   "DB_MouldEditor_HMI_uData_arShotSet{0}_Pressure{4}" : Real = PLC DB_MouldEditor_HMI.uData.arShotSet[0].Pressure[4] AT %DB10.DBD126, 1 s
   "DB_MouldEditor_HMI_uData_arShotSet{0}_Pressure{5}" : Real = PLC DB_MouldEditor_HMI.uData.arShotSet[0].Pressure[5] AT %DB10.DBD130, 1 s
   "DB_MouldEditor_HMI_uData_arShotSet{0}_Pressure{6}" : Real = PLC DB_MouldEditor_HMI.uData.arShotSet[0].Pressure[6] AT %DB10.DBD134, 1 s
   "DB_MouldEditor_HMI_uData_arShotSet{0}_Flow{1}" : Real = PLC DB_MouldEditor_HMI.uData.arShotSet[0].Flow[1] AT %DB10.DBD138, 1 s
   "DB_MouldEditor_HMI_uData_arShotSet{0}_Flow{2}" : Real = PLC DB_MouldEditor_HMI.uData.arShotSet[0].Flow[2] AT %DB10.DBD142, 1 s
   "DB_MouldEditor_HMI_uData_arShotSet{0}_Flow{3}" : Real = PLC DB_MouldEditor_HMI.uData.arShotSet[0].Flow[3] AT %DB10.DBD146, 1 s
   "DB_MouldEditor_HMI_uData_arShotSet{0}_Flow{4}" : Real = PLC DB_MouldEditor_HMI.uData.arShotSet[0].Flow[4] AT %DB10.DBD150, 1 s
   "DB_MouldEditor_HMI_uData_arShotSet{0}_Flow{5}" : Real = PLC DB_MouldEditor_HMI.uData.arShotSet[0].Flow[5] AT %DB10.DBD154, 1 s
   "DB_MouldEditor_HMI_uData_arShotSet{0}_Flow{6}" : Real = PLC DB_MouldEditor_HMI.uData.arShotSet[0].Flow[6] AT %DB10.DBD158, 1 s
   "DB_MouldEditor_HMI_uData_arShotSet{1}_Pressure{1}" : Real = PLC DB_MouldEditor_HMI.uData.arShotSet[1].Pressure[1] AT %DB10.DBD186, 1 s
   "DB_MouldEditor_HMI_uData_arShotSet{1}_Pressure{2}" : Real = PLC DB_MouldEditor_HMI.uData.arShotSet[1].Pressure[2] AT %DB10.DBD190, 1 s
   "DB_MouldEditor_HMI_uData_arShotSet{1}_Pressure{3}" : Real = PLC DB_MouldEditor_HMI.uData.arShotSet[1].Pressure[3] AT %DB10.DBD194, 1 s
   "DB_MouldEditor_HMI_uData_arShotSet{1}_Pressure{4}" : Real = PLC DB_MouldEditor_HMI.uData.arShotSet[1].Pressure[4] AT %DB10.DBD198, 1 s
   "DB_MouldEditor_HMI_uData_arShotSet{1}_Pressure{5}" : Real = PLC DB_MouldEditor_HMI.uData.arShotSet[1].Pressure[5] AT %DB10.DBD202, 1 s
   "DB_MouldEditor_HMI_uData_arShotSet{1}_Pressure{6}" : Real = PLC DB918_ShotResultlast10.FilteredShot[2].Mixingratio[1] AT %DB10.DBD206, 1 s
   "DB_MouldEditor_HMI_uData_arShotSet{1}_Flow{1}" : Real = PLC DB_MouldEditor_HMI.uData.arShotSet[1].Flow[1] AT %DB10.DBD210, 1 s
   "DB_MouldEditor_HMI_uData_arShotSet{1}_Flow{2}" : Real = PLC DB_MouldEditor_HMI.uData.arShotSet[1].Flow[2] AT %DB10.DBD214, 1 s
   "DB_MouldEditor_HMI_uData_arShotSet{1}_Flow{3}" : Real = PLC DB_MouldEditor_HMI.uData.arShotSet[1].Flow[3] AT %DB10.DBD218, 1 s
   "DB_MouldEditor_HMI_uData_arShotSet{1}_Flow{4}" : Real = PLC DB_MouldEditor_HMI.uData.arShotSet[1].Flow[4] AT %DB10.DBD222, 1 s
   "DB_MouldEditor_HMI_uData_arShotSet{1}_Flow{5}" : Real = PLC DB_MouldEditor_HMI.uData.arShotSet[1].Flow[5] AT %DB10.DBD226, 1 s
   "DB_MouldEditor_HMI_uData_arShotSet{1}_Flow{6}" : Real = PLC DB_MouldEditor_HMI.uData.arShotSet[1].Flow[6] AT %DB10.DBD230, 1 s
   "DB_MouldEditor_HMI_uData_arShotSet{2}_Pressure{1}" : Real = PLC DB_MouldEditor_HMI.uData.arShotSet[2].Pressure[1] AT %DB10.DBD258, 1 s
   "DB_MouldEditor_HMI_uData_arShotSet{2}_Pressure{2}" : Real = PLC DB_MouldEditor_HMI.uData.arShotSet[2].Pressure[2] AT %DB10.DBD262, 1 s
   "DB_MouldEditor_HMI_uData_arShotSet{2}_Pressure{3}" : Real = PLC DB_MouldEditor_HMI.uData.arShotSet[2].Pressure[3] AT %DB10.DBD266, 1 s
   "DB_MouldEditor_HMI_uData_arShotSet{2}_Pressure{4}" : Real = PLC DB_MouldEditor_HMI.uData.arShotSet[2].Pressure[4] AT %DB10.DBD270, 1 s
   "DB_MouldEditor_HMI_uData_arShotSet{2}_Pressure{5}" : Real = PLC DB_MouldEditor_HMI.uData.arShotSet[2].Pressure[5] AT %DB10.DBD274, 1 s
   "DB_MouldEditor_HMI_uData_arShotSet{2}_Pressure{6}" : Real = PLC DB_MouldEditor_HMI.uData.arShotSet[2].Pressure[6] AT %DB10.DBD278, 1 s
   "DB_MouldEditor_HMI_uData_arShotSet{2}_Flow{1}" : Real = PLC DB_MouldEditor_HMI.uData.arShotSet[2].Flow[1] AT %DB10.DBD282, 1 s
   "DB_MouldEditor_HMI_uData_arShotSet{2}_Flow{2}" : Real = PLC DB_MouldEditor_HMI.uData.arShotSet[2].Flow[2] AT %DB10.DBD286, 1 s
   "DB_MouldEditor_HMI_uData_arShotSet{2}_Flow{3}" : Real = PLC DB_MouldEditor_HMI.uData.arShotSet[2].Flow[3] AT %DB10.DBD290, 1 s
   "DB_MouldEditor_HMI_uData_arShotSet{2}_Flow{4}" : Real = PLC DB_MouldEditor_HMI.uData.arShotSet[2].Flow[4] AT %DB10.DBD294, 1 s
   "DB_MouldEditor_HMI_uData_arShotSet{2}_Flow{5}" : Real = PLC DB_MouldEditor_HMI.uData.arShotSet[2].Flow[5] AT %DB10.DBD298, 1 s
   "DB_MouldEditor_HMI_uData_arShotSet{2}_Flow{6}" : Real = PLC DB_MouldEditor_HMI.uData.arShotSet[2].Flow[6] AT %DB10.DBD302, 1 s
   "DB_MouldEditor_HMI_uData_arShotSet{3}_Pressure{1}" : Real = PLC DB_MouldEditor_HMI.uData.arShotSet[3].Pressure[1] AT %DB10.DBD330, 1 s
   "DB_MouldEditor_HMI_uData_arShotSet{3}_Pressure{2}" : Real = PLC DB_MouldEditor_HMI.uData.arShotSet[3].Pressure[2] AT %DB10.DBD334, 1 s
   "DB_MouldEditor_HMI_uData_arShotSet{3}_Pressure{3}" : Real = PLC DB_MouldEditor_HMI.uData.arShotSet[3].Pressure[3] AT %DB10.DBD338, 1 s
   "DB_MouldEditor_HMI_uData_arShotSet{3}_Pressure{4}" : Real = PLC DB_MouldEditor_HMI.uData.arShotSet[3].Pressure[4] AT %DB10.DBD342, 1 s
   "DB_MouldEditor_HMI_uData_arShotSet{3}_Pressure{5}" : Real = PLC DB_MouldEditor_HMI.uData.arShotSet[3].Pressure[5] AT %DB10.DBD346, 1 s
   "DB_MouldEditor_HMI_uData_arShotSet{3}_Pressure{6}" : Real = PLC DB_MouldEditor_HMI.uData.arShotSet[3].Pressure[6] AT %DB10.DBD350, 1 s
   "DB_MouldEditor_HMI_uData_arShotSet{3}_Flow{1}" : Real = PLC DB_MouldEditor_HMI.uData.arShotSet[3].Flow[1] AT %DB10.DBD354, 1 s
   "DB_MouldEditor_HMI_uData_arShotSet{3}_Flow{2}" : Real = PLC DB_MouldEditor_HMI.uData.arShotSet[3].Flow[2] AT %DB10.DBD358, 1 s
   "DB_MouldEditor_HMI_uData_arShotSet{3}_Flow{3}" : Real = PLC DB_MouldEditor_HMI.uData.arShotSet[3].Flow[3] AT %DB10.DBD362, 1 s
   "DB_MouldEditor_HMI_uData_arShotSet{3}_Flow{4}" : Real = PLC DB_MouldEditor_HMI.uData.arShotSet[3].Flow[4] AT %DB10.DBD366, 1 s
   "DB_MouldEditor_HMI_uData_arShotSet{3}_Flow{5}" : Real = PLC DB_MouldEditor_HMI.uData.arShotSet[3].Flow[5] AT %DB10.DBD370, 1 s
   "DB_MouldEditor_HMI_uData_arShotSet{3}_Flow{6}" : Real = PLC DB_MouldEditor_HMI.uData.arShotSet[3].Flow[6] AT %DB10.DBD374, 1 s
   "DB_MouldEditor_HMI_uData_arShotSet{4}_Pressure{1}" : Real = PLC DB_MouldEditor_HMI.uData.arShotSet[4].Pressure[1] AT %DB10.DBD402, 1 s
   "DB_MouldEditor_HMI_uData_arShotSet{4}_Pressure{2}" : Real = PLC DB_MouldEditor_HMI.uData.arShotSet[4].Pressure[2] AT %DB10.DBD406, 1 s
   "DB_MouldEditor_HMI_uData_arShotSet{4}_Pressure{3}" : Real = PLC DB_MouldEditor_HMI.uData.arShotSet[4].Pressure[3] AT %DB10.DBD410, 1 s
   "DB_MouldEditor_HMI_uData_arShotSet{4}_Pressure{4}" : Real = PLC DB_MouldEditor_HMI.uData.arShotSet[4].Pressure[4] AT %DB10.DBD414, 1 s
   "DB_MouldEditor_HMI_uData_arShotSet{4}_Pressure{5}" : Real = PLC DB_MouldEditor_HMI.uData.arShotSet[4].Pressure[5] AT %DB10.DBD418, 1 s
   "DB_MouldEditor_HMI_uData_arShotSet{4}_Pressure{6}" : Real = PLC DB_MouldEditor_HMI.uData.arShotSet[4].Pressure[6] AT %DB10.DBD422, 1 s
   "DB_MouldEditor_HMI_uData_arShotSet{4}_Flow{1}" : Real = PLC DB_MouldEditor_HMI.uData.arShotSet[4].Flow[1] AT %DB10.DBD426, 1 s
   "DB_MouldEditor_HMI_uData_arShotSet{4}_Flow{2}" : Real = PLC DB_MouldEditor_HMI.uData.arShotSet[4].Flow[2] AT %DB10.DBD430, 1 s
   "DB_MouldEditor_HMI_uData_arShotSet{4}_Flow{3}" : Real = PLC DB_MouldEditor_HMI.uData.arShotSet[4].Flow[3] AT %DB10.DBD434, 1 s
   "DB_MouldEditor_HMI_uData_arShotSet{4}_Flow{4}" : Real = PLC DB_MouldEditor_HMI.uData.arShotSet[4].Flow[4] AT %DB10.DBD438, 1 s
   "DB_MouldEditor_HMI_uData_arShotSet{4}_Flow{5}" : Real = PLC DB_MouldEditor_HMI.uData.arShotSet[4].Flow[5] AT %DB10.DBD442, 1 s
   "DB_MouldEditor_HMI_uData_arShotSet{4}_Flow{6}" : Real = PLC DB_MouldEditor_HMI.uData.arShotSet[4].Flow[6] AT %DB10.DBD446, 1 s
   "DB_MouldEditor_HMI_uData_arShotSet{5}_Pressure{1}" : Real = PLC DB_MouldEditor_HMI.uData.arShotSet[5].Pressure[1] AT %DB10.DBD474, 1 s
   "DB_MouldEditor_HMI_uData_arShotSet{5}_Pressure{2}" : Real = PLC DB_MouldEditor_HMI.uData.arShotSet[5].Pressure[2] AT %DB10.DBD478, 1 s
   "DB_MouldEditor_HMI_uData_arShotSet{5}_Pressure{3}" : Real = PLC DB_MouldEditor_HMI.uData.arShotSet[5].Pressure[3] AT %DB10.DBD482, 1 s
   "DB_MouldEditor_HMI_uData_arShotSet{5}_Pressure{4}" : Real = PLC DB_MouldEditor_HMI.uData.arShotSet[5].Pressure[4] AT %DB10.DBD486, 1 s
   "DB_MouldEditor_HMI_uData_arShotSet{5}_Pressure{5}" : Real = PLC DB_MouldEditor_HMI.uData.arShotSet[5].Pressure[5] AT %DB10.DBD490, 1 s
   "DB_MouldEditor_HMI_uData_arShotSet{5}_Pressure{6}" : Real = PLC DB_MouldEditor_HMI.uData.arShotSet[5].Pressure[6] AT %DB10.DBD494, 1 s
   "DB_MouldEditor_HMI_uData_arShotSet{5}_Flow{1}" : Real = PLC DB_MouldEditor_HMI.uData.arShotSet[5].Flow[1] AT %DB10.DBD498, 1 s
   "DB_MouldEditor_HMI_uData_arShotSet{5}_Flow{2}" : Real = PLC DB_MouldEditor_HMI.uData.arShotSet[5].Flow[2] AT %DB10.DBD502, 1 s
   "DB_MouldEditor_HMI_uData_arShotSet{5}_Flow{3}" : Real = PLC DB_MouldEditor_HMI.uData.arShotSet[5].Flow[3] AT %DB10.DBD506, 1 s
   "DB_MouldEditor_HMI_uData_arShotSet{5}_Flow{4}" : Real = PLC DB_MouldEditor_HMI.uData.arShotSet[5].Flow[4] AT %DB10.DBD510, 1 s
   "DB_MouldEditor_HMI_uData_arShotSet{5}_Flow{5}" : Real = PLC DB_MouldEditor_HMI.uData.arShotSet[5].Flow[5] AT %DB10.DBD514, 1 s
   "DB_MouldEditor_HMI_uData_arShotSet{5}_Flow{6}" : Real = PLC DB_MouldEditor_HMI.uData.arShotSet[5].Flow[6] AT %DB10.DBD518, 1 s
   "DB_MouldEditor_HMI_uData_arShotSet{6}_Pressure{1}" : Real = PLC DB_MouldEditor_HMI.uData.arShotSet[6].Pressure[1] AT %DB10.DBD546, 1 s
   "DB_MouldEditor_HMI_uData_arShotSet{6}_Pressure{2}" : Real = PLC DB_MouldEditor_HMI.uData.arShotSet[6].Pressure[2] AT %DB10.DBD550, 1 s
   "DB_MouldEditor_HMI_uData_arShotSet{6}_Pressure{3}" : Real = PLC DB_MouldEditor_HMI.uData.arShotSet[6].Pressure[3] AT %DB10.DBD554, 1 s
   "DB_MouldEditor_HMI_uData_arShotSet{6}_Pressure{4}" : Real = PLC DB_MouldEditor_HMI.uData.arShotSet[6].Pressure[4] AT %DB10.DBD558, 1 s
   "DB_MouldEditor_HMI_uData_arShotSet{6}_Pressure{5}" : Real = PLC DB_MouldEditor_HMI.uData.arShotSet[6].Pressure[5] AT %DB10.DBD562, 1 s
   "DB_MouldEditor_HMI_uData_arShotSet{6}_Pressure{6}" : Real = PLC DB_MouldEditor_HMI.uData.arShotSet[6].Pressure[6] AT %DB10.DBD566, 1 s
   "DB_MouldEditor_HMI_uData_arShotSet{6}_Flow{1}" : Real = PLC DB_MouldEditor_HMI.uData.arShotSet[6].Flow[1] AT %DB10.DBD570, 1 s
   "DB_MouldEditor_HMI_uData_arShotSet{6}_Flow{2}" : Real = PLC DB_MouldEditor_HMI.uData.arShotSet[6].Flow[2] AT %DB10.DBD574, 1 s
   "DB_MouldEditor_HMI_uData_arShotSet{6}_Flow{3}" : Real = PLC DB_MouldEditor_HMI.uData.arShotSet[6].Flow[3] AT %DB10.DBD578, 1 s
   "DB_MouldEditor_HMI_uData_arShotSet{6}_Flow{4}" : Real = PLC DB_MouldEditor_HMI.uData.arShotSet[6].Flow[4] AT %DB10.DBD582, 1 s
   "DB_MouldEditor_HMI_uData_arShotSet{6}_Flow{5}" : Real = PLC DB_MouldEditor_HMI.uData.arShotSet[6].Flow[5] AT %DB10.DBD586, 1 s
   "DB_MouldEditor_HMI_uData_arShotSet{6}_Flow{6}" : Real = PLC DB_MouldEditor_HMI.uData.arShotSet[6].Flow[6] AT %DB10.DBD590, 1 s
   "DB_MouldEditor_HMI_uData_arShotSet{7}_Pressure{1}" : Real = PLC DB_MouldEditor_HMI.uData.arShotSet[7].Pressure[1] AT %DB10.DBD618, 1 s
   "DB_MouldEditor_HMI_uData_arShotSet{7}_Pressure{2}" : Real = PLC DB_MouldEditor_HMI.uData.arShotSet[7].Pressure[2] AT %DB10.DBD622, 1 s
   "DB_MouldEditor_HMI_uData_arShotSet{7}_Pressure{3}" : Real = PLC DB_MouldEditor_HMI.uData.arShotSet[7].Pressure[3] AT %DB10.DBD626, 1 s
   "DB_MouldEditor_HMI_uData_arShotSet{7}_Pressure{4}" : Real = PLC DB_MouldEditor_HMI.uData.arShotSet[7].Pressure[4] AT %DB10.DBD630, 1 s
   "DB_MouldEditor_HMI_uData_arShotSet{7}_Pressure{5}" : Real = PLC DB_MouldEditor_HMI.uData.arShotSet[7].Pressure[5] AT %DB10.DBD634, 1 s
   "DB_MouldEditor_HMI_uData_arShotSet{7}_Pressure{6}" : Real = PLC DB_MouldEditor_HMI.uData.arShotSet[7].Pressure[6] AT %DB10.DBD638, 1 s
   "DB_MouldEditor_HMI_uData_arShotSet{7}_Flow{1}" : Real = PLC DB_MouldEditor_HMI.uData.arShotSet[7].Flow[1] AT %DB10.DBD642, 1 s
   "DB_MouldEditor_HMI_uData_arShotSet{7}_Flow{2}" : Real = PLC DB_MouldEditor_HMI.uData.arShotSet[7].Flow[2] AT %DB10.DBD646, 1 s
   "DB_MouldEditor_HMI_uData_arShotSet{7}_Flow{3}" : Real = PLC DB_MouldEditor_HMI.uData.arShotSet[7].Flow[3] AT %DB10.DBD650, 1 s
   "DB_MouldEditor_HMI_uData_arShotSet{7}_Flow{4}" : Real = PLC DB_MouldEditor_HMI.uData.arShotSet[7].Flow[4] AT %DB10.DBD654, 1 s
   "DB_MouldEditor_HMI_uData_arShotSet{7}_Flow{5}" : Real = PLC DB_MouldEditor_HMI.uData.arShotSet[7].Flow[5] AT %DB10.DBD658, 1 s
   "DB_MouldEditor_HMI_uData_arShotSet{7}_Flow{6}" : Real = PLC DB_MouldEditor_HMI.uData.arShotSet[7].Flow[6] AT %DB10.DBD662, 1 s
   "DB_MouldEditor_HMI_uData_arShotSet{8}_Pressure{1}" : Real = PLC DB_MouldEditor_HMI.uData.arShotSet[8].Pressure[1] AT %DB10.DBD690, 1 s
   "DB_MouldEditor_HMI_uData_arShotSet{8}_Pressure{2}" : Real = PLC DB_MouldEditor_HMI.uData.arShotSet[8].Pressure[2] AT %DB10.DBD694, 1 s
   "DB_MouldEditor_HMI_uData_arShotSet{8}_Pressure{3}" : Real = PLC DB_MouldEditor_HMI.uData.arShotSet[8].Pressure[3] AT %DB10.DBD698, 1 s
   "DB_MouldEditor_HMI_uData_arShotSet{8}_Pressure{4}" : Real = PLC DB_MouldEditor_HMI.uData.arShotSet[8].Pressure[4] AT %DB10.DBD702, 1 s
   "DB_MouldEditor_HMI_uData_arShotSet{8}_Pressure{5}" : Real = PLC DB_MouldEditor_HMI.uData.arShotSet[8].Pressure[5] AT %DB10.DBD706, 1 s
   "DB_MouldEditor_HMI_uData_arShotSet{8}_Pressure{6}" : Real = PLC DB_MouldEditor_HMI.uData.arShotSet[8].Pressure[6] AT %DB10.DBD710, 1 s
   "DB_MouldEditor_HMI_uData_arShotSet{8}_Flow{1}" : Real = PLC DB_MouldEditor_HMI.uData.arShotSet[8].Flow[1] AT %DB10.DBD714, 1 s
   "DB_MouldEditor_HMI_uData_arShotSet{8}_Flow{2}" : Real = PLC DB_MouldEditor_HMI.uData.arShotSet[8].Flow[2] AT %DB10.DBD718, 1 s
   "DB_MouldEditor_HMI_uData_arShotSet{8}_Flow{3}" : Real = PLC DB_MouldEditor_HMI.uData.arShotSet[8].Flow[3] AT %DB10.DBD722, 1 s
   "DB_MouldEditor_HMI_uData_arShotSet{8}_Flow{4}" : Real = PLC DB_MouldEditor_HMI.uData.arShotSet[8].Flow[4] AT %DB10.DBD726, 1 s
   "DB_MouldEditor_HMI_uData_arShotSet{8}_Flow{5}" : Real = PLC DB_MouldEditor_HMI.uData.arShotSet[8].Flow[5] AT %DB10.DBD730, 1 s
   "DB_MouldEditor_HMI_uData_arShotSet{8}_Flow{6}" : Real = PLC DB_MouldEditor_HMI.uData.arShotSet[8].Flow[6] AT %DB10.DBD734, 1 s
   "DB930_Tools_Tool{1}_tool_name" : String[20] = PLC DB930_Tools.Tool[1].tool_name AT %DB930.DBX44.0, 1 s
   "DB930_Tools_Tool{2}_tool_name" : String[20] = PLC DB930_Tools.Tool[2].tool_name AT %DB930.DBX78.0, 1 s
   "DB930_Tools_Tool{3}_tool_name" : String[20] = PLC DB930_Tools.Tool[3].tool_name AT %DB930.DBX112.0, 1 s
   "DB930_Tools_Tool{4}_tool_name" : String[20] = PLC DB930_Tools.Tool[4].tool_name AT %DB930.DBX146.0, 1 s
   "DB930_Tools_Tool{5}_tool_name" : String[20] = PLC DB930_Tools.Tool[5].tool_name AT %DB930.DBX180.0, 1 s
   "DB930_Tools_Tool{6}_tool_name" : String[20] = PLC DB930_Tools.Tool[6].tool_name AT %DB930.DBX214.0, 1 s
   "DB930_Tools_Tool{7}_tool_name" : String[20] = PLC DB930_Tools.Tool[7].tool_name AT %DB930.DBX248.0, 1 s
   "DB930_Tools_Tool{8}_tool_name" : String[20] = PLC DB930_Tools.Tool[8].tool_name AT %DB930.DBX282.0, 1 s
   "DB930_Tools_Tool{9}_tool_name" : String[20] = PLC DB930_Tools.Tool[9].tool_name AT %DB930.DBX316.0, 1 s
   "DB930_Tools_Tool{10}_tool_name" : String[20] = PLC DB930_Tools.Tool[10].tool_name AT %DB930.DBX350.0, 1 s
   "DB930_Tools_Tool{11}_tool_name" : String[20] = PLC DB930_Tools.Tool[11].tool_name AT %DB930.DBX384.0, 1 s
   "DB930_Tools_Tool{12}_tool_name" : String[20] = PLC DB930_Tools.Tool[12].tool_name AT %DB930.DBX418.0, 1 s
   "DB930_Tools_Tool{13}_tool_name" : String[20] = PLC DB930_Tools.Tool[13].tool_name AT %DB930.DBX452.0, 1 s
   "DB930_Tools_Tool{14}_tool_name" : String[20] = PLC DB930_Tools.Tool[14].tool_name AT %DB930.DBX486.0, 1 s
   "DB930_Tools_Tool{15}_tool_name" : String[20] = PLC DB930_Tools.Tool[15].tool_name AT %DB930.DBX520.0, 1 s
   "DB930_Tools_Tool{16}_tool_name" : String[20] = PLC DB930_Tools.Tool[16].tool_name AT %DB930.DBX554.0, 1 s
   "DB930_Tools_Tool{17}_tool_name" : String[20] = PLC DB930_Tools.Tool[17].tool_name AT %DB930.DBX588.0, 1 s
   "DB930_Tools_Tool{18}_tool_name" : String[20] = PLC DB930_Tools.Tool[18].tool_name AT %DB930.DBX622.0, 1 s
   "DB930_Tools_Tool{19}_tool_name" : String[20] = PLC DB930_Tools.Tool[19].tool_name AT %DB930.DBX656.0, 1 s
   "DB930_Tools_Tool{20}_tool_name" : String[20] = PLC DB930_Tools.Tool[20].tool_name AT %DB930.DBX690.0, 1 s
   "DB930_Tools_Tool{21}_tool_name" : String[20] = PLC DB930_Tools.Tool[21].tool_name AT %DB930.DBX724.0, 1 s
   "DB930_Tools_Tool{22}_tool_name" : String[20] = PLC DB930_Tools.Tool[22].tool_name AT %DB930.DBX758.0, 1 s
   "DB930_Tools_Tool{23}_tool_name" : String[20] = PLC DB930_Tools.Tool[23].tool_name AT %DB930.DBX792.0, 1 s
   "DB930_Tools_Tool{24}_tool_name" : String[20] = PLC DB930_Tools.Tool[24].tool_name AT %DB930.DBX826.0, 1 s
   "DB930_Tools_Tool{25}_tool_name" : String[20] = PLC DB930_Tools.Tool[25].tool_name AT %DB930.DBX860.0, 1 s
   "DB930_Tools_Tool{26}_tool_name" : String[20] = PLC DB930_Tools.Tool[26].tool_name AT %DB930.DBX894.0, 1 s
   "DB930_Tools_Tool{27}_tool_name" : String[20] = PLC DB930_Tools.Tool[27].tool_name AT %DB930.DBX928.0, 1 s
   "DB930_Tools_Tool{28}_tool_name" : String[20] = PLC DB930_Tools.Tool[28].tool_name AT %DB930.DBX962.0, 1 s
   "DB930_Tools_Tool{29}_tool_name" : String[20] = PLC DB930_Tools.Tool[29].tool_name AT %DB930.DBX996.0, 1 s
   "DB930_Tools_Tool{30}_tool_name" : String[20] = PLC DB930_Tools.Tool[30].tool_name AT %DB930.DBX1030.0, 1 s
   "DB930_Tools_Tool{31}_tool_name" : String[20] = PLC DB930_Tools.Tool[31].tool_name AT %DB930.DBX1064.0, 1 s
   "DB930_Tools_Tool{32}_tool_name" : String[20] = PLC DB930_Tools.Tool[32].tool_name AT %DB930.DBX1098.0, 1 s
   "DB930_Tools_Tool{33}_tool_name" : String[20] = PLC DB930_Tools.Tool[33].tool_name AT %DB930.DBX1132.0, 1 s
   "DB930_Tools_Tool{34}_tool_name" : String[20] = PLC DB930_Tools.Tool[34].tool_name AT %DB930.DBX1166.0, 1 s
   "DB930_Tools_Tool{35}_tool_name" : String[20] = PLC DB930_Tools.Tool[35].tool_name AT %DB930.DBX1200.0, 1 s
   "DB930_Tools_Tool{36}_tool_name" : String[20] = PLC DB930_Tools.Tool[36].tool_name AT %DB930.DBX1234.0, 1 s
   "DB930_Tools_Tool{37}_tool_name" : String[20] = PLC DB930_Tools.Tool[37].tool_name AT %DB930.DBX1268.0, 1 s
   "DB930_Tools_Tool{38}_tool_name" : String[20] = PLC DB930_Tools.Tool[38].tool_name AT %DB930.DBX1302.0, 1 s
   "DB930_Tools_Tool{39}_tool_name" : String[20] = PLC DB930_Tools.Tool[39].tool_name AT %DB930.DBX1336.0, 1 s
   "DB930_Tools_Tool{40}_tool_name" : String[20] = PLC DB930_Tools.Tool[40].tool_name AT %DB930.DBX1370.0, 1 s
   "DB930_Tools_Tool{41}_tool_name" : String[20] = PLC DB930_Tools.Tool[41].tool_name AT %DB930.DBX1404.0, 1 s
   "DB930_Tools_Tool{42}_tool_name" : String[20] = PLC DB930_Tools.Tool[42].tool_name AT %DB930.DBX1438.0, 1 s
   "DB930_Tools_Tool{43}_tool_name" : String[20] = PLC DB930_Tools.Tool[43].tool_name AT %DB930.DBX1472.0, 1 s
   "DB930_Tools_Tool{44}_tool_name" : String[20] = PLC DB930_Tools.Tool[44].tool_name AT %DB930.DBX1506.0, 1 s
   "DB930_Tools_Tool{45}_tool_name" : String[20] = PLC DB930_Tools.Tool[45].tool_name AT %DB930.DBX1540.0, 1 s
   "DB930_Tools_Tool{46}_tool_name" : String[20] = PLC DB930_Tools.Tool[46].tool_name AT %DB930.DBX1574.0, 1 s
   "DB930_Tools_Tool{47}_tool_name" : String[20] = PLC DB930_Tools.Tool[47].tool_name AT %DB930.DBX1608.0, 1 s
   "DB930_Tools_Tool{48}_tool_name" : String[20] = PLC DB930_Tools.Tool[48].tool_name AT %DB930.DBX1642.0, 1 s
   "DB930_Tools_Tool{49}_tool_name" : String[20] = PLC DB930_Tools.Tool[49].tool_name AT %DB930.DBX1676.0, 1 s
   "DB930_Tools_Tool{50}_tool_name" : String[20] = PLC DB930_Tools.Tool[50].tool_name AT %DB930.DBX1710.0, 1 s
   "DB930_Tools_Tool{51}_tool_name" : String[20] = PLC DB930_Tools.Tool[51].tool_name AT %DB930.DBX1744.0, 1 s
   "DB930_Tools_Tool{52}_tool_name" : String[20] = PLC DB930_Tools.Tool[52].tool_name AT %DB930.DBX1778.0, 1 s
   "DB930_Tools_Tool{53}_tool_name" : String[20] = PLC DB930_Tools.Tool[53].tool_name AT %DB930.DBX1812.0, 1 s
   "DB930_Tools_Tool{54}_tool_name" : String[20] = PLC DB930_Tools.Tool[54].tool_name AT %DB930.DBX1846.0, 1 s
   "DB930_Tools_Tool{55}_tool_name" : String[20] = PLC DB930_Tools.Tool[55].tool_name AT %DB930.DBX1880.0, 1 s
   "DB930_Tools_Tool{56}_tool_name" : String[20] = PLC DB930_Tools.Tool[56].tool_name AT %DB930.DBX1914.0, 1 s
   "DB930_Tools_Tool{57}_tool_name" : String[20] = PLC DB930_Tools.Tool[57].tool_name AT %DB930.DBX1948.0, 1 s
   "DB930_Tools_Tool{58}_tool_name" : String[20] = PLC DB930_Tools.Tool[58].tool_name AT %DB930.DBX1982.0, 1 s
   "DB930_Tools_Tool{59}_tool_name" : String[20] = PLC DB930_Tools.Tool[59].tool_name AT %DB930.DBX2016.0, 1 s
   "DB930_Tools_Tool{60}_tool_name" : String[20] = PLC DB930_Tools.Tool[60].tool_name AT %DB930.DBX2050.0, 1 s
   "DB_MouldEditor_HMI_uData_sSelected_sPS_arFlow{0}" : Real = PLC DB_MouldEditor_HMI.uData.sSelected.sPS.arFlow[0] AT %DB10.DBD4, 1 s
   "DB_MouldEditor_HMI_uData_sSelected_sPS_arRatio{0}" : Real = PLC DB_MouldEditor_HMI.uData.sSelected.sPS.arRatio[0] AT %DB10.DBD32, 1 s
   "DB_MouldEditor_HMI_uData_sSelected_sPS_arPressure{0}" : Real = PLC DB_MouldEditor_HMI.uData.sSelected.sPS.arPressure[0] AT %DB10.DBD60, 1 s
   "DB_MouldEditor_HMI_uData_sSelected_sPS_2PoinMovement_Comp01" : Bool = PLC DB_MouldEditor_HMI.uData.sSelected.sPS.2PoinMovement_Comp01 AT %DB10.DBX90.0, 1 s
   "DB_MouldEditor_HMI_uData_sSelected_sPS_2PoinMovement_Comp02" : Bool = PLC DB_MouldEditor_HMI.uData.sSelected.sPS.2PoinMovement_Comp02 AT %DB10.DBX90.1, 1 s
   "DB_MouldEditor_HMI_uData_sSelected_sPS_2PoinMovement_Comp03" : Bool = PLC DB_MouldEditor_HMI.uData.sSelected.sPS.2PoinMovement_Comp03 AT %DB10.DBX90.2, 1 s
   "DB_MouldEditor_HMI_uData_sSelected_sPS_2PoinMovement_Comp04" : Bool = PLC DB_MouldEditor_HMI.uData.sSelected.sPS.2PoinMovement_Comp04 AT %DB10.DBX90.3, 1 s
   "DB_MouldEditor_HMI_uData_sSelected_sPS_2PoinMovement_Comp05" : Bool = PLC DB_MouldEditor_HMI.uData.sSelected.sPS.2PoinMovement_Comp05 AT %DB10.DBX90.4, 1 s
   "DB_MouldEditor_HMI_uData_sSelected_sPS_2PoinMovement_Comp06" : Bool = PLC DB_MouldEditor_HMI.uData.sSelected.sPS.2PoinMovement_Comp06 AT %DB10.DBX90.5, 1 s
   "DB930_Tools_Tool{61}_tool_name" : String[20] = PLC DB930_Tools.Tool[61].tool_name AT %DB930.DBX2084.0, 1 s
   "DB930_Tools_Tool{62}_tool_name" : String[20] = PLC DB930_Tools.Tool[62].tool_name AT %DB930.DBX2118.0, 1 s
   "DB930_Tools_Tool{63}_tool_name" : String[20] = PLC DB930_Tools.Tool[63].tool_name AT %DB930.DBX2152.0, 1 s
   "DB930_Tools_Tool{64}_tool_name" : String[20] = PLC DB930_Tools.Tool[64].tool_name AT %DB930.DBX2186.0, 1 s
   "DB930_Tools_Tool{65}_tool_name" : String[20] = PLC DB930_Tools.Tool[65].tool_name AT %DB930.DBX2220.0, 1 s
   "DB930_Tools_Tool{66}_tool_name" : String[20] = PLC DB930_Tools.Tool[66].tool_name AT %DB930.DBX2254.0, 1 s
   "DB930_Tools_Tool{67}_tool_name" : String[20] = PLC DB930_Tools.Tool[67].tool_name AT %DB930.DBX2288.0, 1 s
   "DB930_Tools_Tool{68}_tool_name" : String[20] = PLC DB930_Tools.Tool[68].tool_name AT %DB930.DBX2322.0, 1 s
   "DB930_Tools_Tool{69}_tool_name" : String[20] = PLC DB930_Tools.Tool[69].tool_name AT %DB930.DBX2356.0, 1 s
   "DB930_Tools_Tool{70}_tool_name" : String[20] = PLC DB930_Tools.Tool[70].tool_name AT %DB930.DBX2390.0, 1 s
   "DB930_Tools_Tool{71}_tool_name" : String[20] = PLC DB930_Tools.Tool[71].tool_name AT %DB930.DBX2424.0, 1 s
   "DB930_Tools_Tool{72}_tool_name" : String[20] = PLC DB930_Tools.Tool[72].tool_name AT %DB930.DBX2458.0, 1 s
   "DB930_Tools_Tool{73}_tool_name" : String[20] = PLC DB930_Tools.Tool[73].tool_name AT %DB930.DBX2492.0, 1 s
   "DB930_Tools_Tool{74}_tool_name" : String[20] = PLC DB930_Tools.Tool[74].tool_name AT %DB930.DBX2526.0, 1 s
   "DB930_Tools_Tool{75}_tool_name" : String[20] = PLC DB930_Tools.Tool[75].tool_name AT %DB930.DBX2560.0, 1 s
   "DB930_Tools_Tool{76}_tool_name" : String[20] = PLC DB930_Tools.Tool[76].tool_name AT %DB930.DBX2594.0, 1 s
   "DB930_Tools_Tool{77}_tool_name" : String[20] = PLC DB930_Tools.Tool[77].tool_name AT %DB930.DBX2628.0, 1 s
   "DB930_Tools_Tool{78}_tool_name" : String[20] = PLC DB930_Tools.Tool[78].tool_name AT %DB930.DBX2662.0, 1 s
   "DB930_Tools_Tool{79}_tool_name" : String[20] = PLC DB930_Tools.Tool[79].tool_name AT %DB930.DBX2696.0, 1 s
   "DB930_Tools_Tool{80}_tool_name" : String[20] = PLC DB930_Tools.Tool[80].tool_name AT %DB930.DBX2730.0, 1 s
   "DB930_Tools_Tool{81}_tool_name" : String[20] = PLC DB930_Tools.Tool[81].tool_name AT %DB930.DBX2764.0, 1 s
   "DB930_Tools_Tool{82}_tool_name" : String[20] = PLC DB930_Tools.Tool[82].tool_name AT %DB930.DBX2798.0, 1 s
   "DB930_Tools_Tool{83}_tool_name" : String[20] = PLC DB930_Tools.Tool[83].tool_name AT %DB930.DBX2832.0, 1 s
   "DB930_Tools_Tool{84}_tool_name" : String[20] = PLC DB930_Tools.Tool[84].tool_name AT %DB930.DBX2866.0, 1 s
   "DB930_Tools_Tool{85}_tool_name" : String[20] = PLC DB930_Tools.Tool[85].tool_name AT %DB930.DBX2900.0, 1 s
   "DB930_Tools_Tool{86}_tool_name" : String[20] = PLC DB930_Tools.Tool[86].tool_name AT %DB930.DBX2934.0, 1 s
   "DB930_Tools_Tool{87}_tool_name" : String[20] = PLC DB930_Tools.Tool[87].tool_name AT %DB930.DBX2968.0, 1 s
   "DB930_Tools_Tool{88}_tool_name" : String[20] = PLC DB930_Tools.Tool[88].tool_name AT %DB930.DBX3002.0, 1 s
   "DB930_Tools_Tool{89}_tool_name" : String[20] = PLC DB930_Tools.Tool[89].tool_name AT %DB930.DBX3036.0, 1 s
   "DB930_Tools_Tool{90}_tool_name" : String[20] = PLC DB930_Tools.Tool[90].tool_name AT %DB930.DBX3070.0, 1 s
   "DB930_Tools_Tool{91}_tool_name" : String[20] = PLC DB930_Tools.Tool[91].tool_name AT %DB930.DBX3104.0, 1 s
   "DB930_Tools_Tool{92}_tool_name" : String[20] = PLC DB930_Tools.Tool[92].tool_name AT %DB930.DBX3138.0, 1 s
   "DB930_Tools_Tool{93}_tool_name" : String[20] = PLC DB930_Tools.Tool[93].tool_name AT %DB930.DBX3172.0, 1 s
   "DB930_Tools_Tool{94}_tool_name" : String[20] = PLC DB930_Tools.Tool[94].tool_name AT %DB930.DBX3206.0, 1 s
   "DB930_Tools_Tool{95}_tool_name" : String[20] = PLC DB930_Tools.Tool[95].tool_name AT %DB930.DBX3240.0, 1 s
   "DB930_Tools_Tool{96}_tool_name" : String[20] = PLC DB930_Tools.Tool[96].tool_name AT %DB930.DBX3274.0, 1 s
   "DB930_Tools_Tool{97}_tool_name" : String[20] = PLC DB930_Tools.Tool[97].tool_name AT %DB930.DBX3308.0, 1 s
   "DB930_Tools_Tool{98}_tool_name" : String[20] = PLC DB930_Tools.Tool[98].tool_name AT %DB930.DBX3342.0, 1 s
   "DB930_Tools_Tool{99}_tool_name" : String[20] = PLC DB930_Tools.Tool[99].tool_name AT %DB930.DBX3376.0, 1 s
   "DB930_Tools_Tool{100}_tool_name" : String[20] = PLC DB930_Tools.Tool[100].tool_name AT %DB930.DBX3410.0, 1 s
   "DB930_Tools_Tool{101}_tool_name" : String[20] = PLC DB930_Tools.Tool[101].tool_name AT %DB930.DBX3444.0, 1 s
   "DB930_Tools_Tool{102}_tool_name" : String[20] = PLC DB930_Tools.Tool[102].tool_name AT %DB930.DBX3478.0, 1 s
   "DB930_Tools_Tool{103}_tool_name" : String[20] = PLC DB930_Tools.Tool[103].tool_name AT %DB930.DBX3512.0, 1 s
   "DB930_Tools_Tool{104}_tool_name" : String[20] = PLC DB930_Tools.Tool[104].tool_name AT %DB930.DBX3546.0, 1 s
   "DB930_Tools_Tool{105}_tool_name" : String[20] = PLC DB930_Tools.Tool[105].tool_name AT %DB930.DBX3580.0, 1 s
   "DB930_Tools_Tool{106}_tool_name" : String[20] = PLC DB930_Tools.Tool[106].tool_name AT %DB930.DBX3614.0, 1 s
   "DB930_Tools_Tool{107}_tool_name" : String[20] = PLC DB930_Tools.Tool[107].tool_name AT %DB930.DBX3648.0, 1 s
   "DB930_Tools_Tool{108}_tool_name" : String[20] = PLC DB930_Tools.Tool[108].tool_name AT %DB930.DBX3682.0, 1 s
   "DB930_Tools_Tool{109}_tool_name" : String[20] = PLC DB930_Tools.Tool[109].tool_name AT %DB930.DBX3716.0, 1 s
   "DB930_Tools_Tool{110}_tool_name" : String[20] = PLC DB930_Tools.Tool[110].tool_name AT %DB930.DBX3750.0, 1 s
   "DB930_Tools_Tool{111}_tool_name" : String[20] = PLC DB930_Tools.Tool[111].tool_name AT %DB930.DBX3784.0, 1 s
   "DB930_Tools_Tool{112}_tool_name" : String[20] = PLC DB930_Tools.Tool[112].tool_name AT %DB930.DBX3818.0, 1 s
   "DB930_Tools_Tool{113}_tool_name" : String[20] = PLC DB930_Tools.Tool[113].tool_name AT %DB930.DBX3852.0, 1 s
   "DB930_Tools_Tool{114}_tool_name" : String[20] = PLC DB930_Tools.Tool[114].tool_name AT %DB930.DBX3886.0, 1 s
   "DB930_Tools_Tool{115}_tool_name" : String[20] = PLC DB930_Tools.Tool[115].tool_name AT %DB930.DBX3920.0, 1 s
   "DB930_Tools_Tool{116}_tool_name" : String[20] = PLC DB930_Tools.Tool[116].tool_name AT %DB930.DBX3954.0, 1 s
   "DB930_Tools_Tool{117}_tool_name" : String[20] = PLC DB930_Tools.Tool[117].tool_name AT %DB930.DBX3988.0, 1 s
   "DB930_Tools_Tool{118}_tool_name" : String[20] = PLC DB930_Tools.Tool[118].tool_name AT %DB930.DBX4022.0, 1 s
   "DB930_Tools_Tool{119}_tool_name" : String[20] = PLC DB930_Tools.Tool[119].tool_name AT %DB930.DBX4056.0, 1 s
   "DB930_Tools_Tool{120}_tool_name" : String[20] = PLC DB930_Tools.Tool[120].tool_name AT %DB930.DBX4090.0, 1 s
   "DB930_Tools_Tool{121}_tool_name" : String[20] = PLC DB930_Tools.Tool[121].tool_name AT %DB930.DBX4124.0, 1 s
   "DB930_Tools_Tool{122}_tool_name" : String[20] = PLC DB930_Tools.Tool[122].tool_name AT %DB930.DBX4158.0, 1 s
   "DB930_Tools_Tool{123}_tool_name" : String[20] = PLC DB930_Tools.Tool[123].tool_name AT %DB930.DBX4192.0, 1 s
   "DB930_Tools_Tool{124}_tool_name" : String[20] = PLC DB930_Tools.Tool[124].tool_name AT %DB930.DBX4226.0, 1 s
   "DB930_Tools_Tool{125}_tool_name" : String[20] = PLC DB930_Tools.Tool[125].tool_name AT %DB930.DBX4260.0, 1 s
   "DB930_Tools_Tool{126}_tool_name" : String[20] = PLC DB930_Tools.Tool[126].tool_name AT %DB930.DBX4294.0, 1 s
   "DB930_Tools_Tool{127}_tool_name" : String[20] = PLC DB930_Tools.Tool[127].tool_name AT %DB930.DBX4328.0, 1 s
   "DB930_Tools_Tool{128}_tool_name" : String[20] = PLC DB930_Tools.Tool[128].tool_name AT %DB930.DBX4362.0, 1 s
   "DB930_Tools_Tool{129}_tool_name" : String[20] = PLC DB930_Tools.Tool[129].tool_name AT %DB930.DBX4396.0, 1 s
   "DB930_Tools_Tool{130}_tool_name" : String[20] = PLC DB930_Tools.Tool[130].tool_name AT %DB930.DBX4430.0, 1 s
   "DB930_Tools_Tool{131}_tool_name" : String[20] = PLC DB930_Tools.Tool[131].tool_name AT %DB930.DBX4464.0, 1 s
   "DB930_Tools_Tool{132}_tool_name" : String[20] = PLC DB930_Tools.Tool[132].tool_name AT %DB930.DBX4498.0, 1 s
   "DB930_Tools_Tool{133}_tool_name" : String[20] = PLC DB930_Tools.Tool[133].tool_name AT %DB930.DBX4532.0, 1 s
   "DB930_Tools_Tool{134}_tool_name" : String[20] = PLC DB930_Tools.Tool[134].tool_name AT %DB930.DBX4566.0, 1 s
   "DB930_Tools_Tool{135}_tool_name" : String[20] = PLC DB930_Tools.Tool[135].tool_name AT %DB930.DBX4600.0, 1 s
   "DB930_Tools_Tool{136}_tool_name" : String[20] = PLC PN_Mixinghead.Mixinghead[0].DüseBypass[2].Visualisierung.PolarityBypass AT %DB930.DBX4634.0, 1 s
   "DB930_Tools_Tool{137}_tool_name" : String[20] = PLC DB930_Tools.Tool[137].tool_name AT %DB930.DBX4668.0, 1 s
   "DB930_Tools_Tool{138}_tool_name" : String[20] = PLC DB930_Tools.Tool[138].tool_name AT %DB930.DBX4702.0, 1 s
   "DB930_Tools_Tool{139}_tool_name" : String[20] = PLC DB930_Tools.Tool[139].tool_name AT %DB930.DBX4736.0, 1 s
   "DB930_Tools_Tool{140}_tool_name" : String[20] = PLC DB930_Tools.Tool[140].tool_name AT %DB930.DBX4770.0, 1 s
   "DB930_Tools_Tool{141}_tool_name" : String[20] = PLC DB930_Tools.Tool[141].tool_name AT %DB930.DBX4804.0, 1 s
   "DB930_Tools_Tool{142}_tool_name" : String[20] = PLC DB930_Tools.Tool[142].tool_name AT %DB930.DBX4838.0, 1 s
   "DB930_Tools_Tool{143}_tool_name" : String[20] = PLC DB930_Tools.Tool[143].tool_name AT %DB930.DBX4872.0, 1 s
   "DB930_Tools_Tool{144}_tool_name" : String[20] = PLC DB930_Tools.Tool[144].tool_name AT %DB930.DBX4906.0, 1 s
   "DB930_Tools_Tool{145}_tool_name" : String[20] = PLC DB930_Tools.Tool[145].tool_name AT %DB930.DBX4940.0, 1 s
   "DB930_Tools_Tool{146}_tool_name" : String[20] = PLC DB930_Tools.Tool[146].tool_name AT %DB930.DBX4974.0, 1 s
   "DB930_Tools_Tool{147}_tool_name" : String[20] = PLC DB930_Tools.Tool[147].tool_name AT %DB930.DBX5008.0, 1 s
   "DB930_Tools_Tool{148}_tool_name" : String[20] = PLC DB930_Tools.Tool[148].tool_name AT %DB930.DBX5042.0, 1 s
   "DB930_Tools_Tool{149}_tool_name" : String[20] = PLC DB930_Tools.Tool[149].tool_name AT %DB930.DBX5076.0, 1 s
   "DB930_Tools_Tool{150}_tool_name" : String[20] = PLC DB930_Tools.Tool[150].tool_name AT %DB930.DBX5110.0, 1 s
   "DB930_Tools_Tool{151}_tool_name" : String[20] = PLC DB930_Tools.Tool[151].tool_name AT %DB930.DBX5144.0, 1 s
   "DB930_Tools_Tool{152}_tool_name" : String[20] = PLC DB930_Tools.Tool[152].tool_name AT %DB930.DBX5178.0, 1 s
   "DB930_Tools_Tool{153}_tool_name" : String[20] = PLC DB930_Tools.Tool[153].tool_name AT %DB930.DBX5212.0, 1 s
   "DB930_Tools_Tool{154}_tool_name" : String[20] = PLC DB930_Tools.Tool[154].tool_name AT %DB930.DBX5246.0, 1 s
   "DB930_Tools_Tool{155}_tool_name" : String[20] = PLC DB930_Tools.Tool[155].tool_name AT %DB930.DBX5280.0, 1 s
   "DB930_Tools_Tool{156}_tool_name" : String[20] = PLC DB930_Tools.Tool[156].tool_name AT %DB930.DBX5314.0, 1 s
   "DB930_Tools_Tool{157}_tool_name" : String[20] = PLC DB930_Tools.Tool[157].tool_name AT %DB930.DBX5348.0, 1 s
   "DB930_Tools_Tool{158}_tool_name" : String[20] = PLC DB930_Tools.Tool[158].tool_name AT %DB930.DBX5382.0, 1 s
   "DB930_Tools_Tool{159}_tool_name" : String[20] = PLC DB930_Tools.Tool[159].tool_name AT %DB930.DBX5416.0, 1 s
   "DB930_Tools_Tool{160}_tool_name" : String[20] = PLC DB930_Tools.Tool[160].tool_name AT %DB930.DBX5450.0, 1 s
   "DB930_Tools_Tool{161}_tool_name" : String[20] = PLC DB930_Tools.Tool[161].tool_name AT %DB930.DBX5484.0, 1 s
   "DB930_Tools_Tool{162}_tool_name" : String[20] = PLC DB930_Tools.Tool[162].tool_name AT %DB930.DBX5518.0, 1 s
   "DB930_Tools_Tool{163}_tool_name" : String[20] = PLC DB930_Tools.Tool[163].tool_name AT %DB930.DBX5552.0, 1 s
   "DB930_Tools_Tool{164}_tool_name" : String[20] = PLC DB930_Tools.Tool[164].tool_name AT %DB930.DBX5586.0, 1 s
   "DB930_Tools_Tool{165}_tool_name" : String[20] = PLC DB930_Tools.Tool[165].tool_name AT %DB930.DBX5620.0, 1 s
   "DB930_Tools_Tool{166}_tool_name" : String[20] = PLC DB930_Tools.Tool[166].tool_name AT %DB930.DBX5654.0, 1 s
   "DB930_Tools_Tool{167}_tool_name" : String[20] = PLC DB930_Tools.Tool[167].tool_name AT %DB930.DBX5688.0, 1 s
   "DB930_Tools_Tool{168}_tool_name" : String[20] = PLC DB930_Tools.Tool[168].tool_name AT %DB930.DBX5722.0, 1 s
   "DB930_Tools_Tool{169}_tool_name" : String[20] = PLC DB930_Tools.Tool[169].tool_name AT %DB930.DBX5756.0, 1 s
   "DB930_Tools_Tool{170}_tool_name" : String[20] = PLC DB930_Tools.Tool[170].tool_name AT %DB930.DBX5790.0, 1 s
   "DB930_Tools_Tool{171}_tool_name" : String[20] = PLC DB930_Tools.Tool[171].tool_name AT %DB930.DBX5824.0, 1 s
   "DB930_Tools_Tool{172}_tool_name" : String[20] = PLC DB930_Tools.Tool[172].tool_name AT %DB930.DBX5858.0, 1 s
   "DB930_Tools_Tool{173}_tool_name" : String[20] = PLC DB930_Tools.Tool[173].tool_name AT %DB930.DBX5892.0, 1 s
   "DB930_Tools_Tool{174}_tool_name" : String[20] = PLC DB930_Tools.Tool[174].tool_name AT %DB930.DBX5926.0, 1 s
   "DB930_Tools_Tool{175}_tool_name" : String[20] = PLC DB930_Tools.Tool[175].tool_name AT %DB930.DBX5960.0, 1 s
   "DB930_Tools_Tool{176}_tool_name" : String[20] = PLC DB930_Tools.Tool[176].tool_name AT %DB930.DBX5994.0, 1 s
   "DB930_Tools_Tool{177}_tool_name" : String[20] = PLC DB930_Tools.Tool[177].tool_name AT %DB930.DBX6028.0, 1 s
   "DB930_Tools_Tool{178}_tool_name" : String[20] = PLC DB930_Tools.Tool[178].tool_name AT %DB930.DBX6062.0, 1 s
   "DB930_Tools_Tool{179}_tool_name" : String[20] = PLC DB930_Tools.Tool[179].tool_name AT %DB930.DBX6096.0, 1 s
   "DB930_Tools_Tool{180}_tool_name" : String[20] = PLC DB930_Tools.Tool[180].tool_name AT %DB930.DBX6130.0, 1 s
   "DB930_Tools_Tool{181}_tool_name" : String[20] = PLC DB930_Tools.Tool[181].tool_name AT %DB930.DBX6164.0, 1 s
   "DB930_Tools_Tool{182}_tool_name" : String[20] = PLC DB930_Tools.Tool[182].tool_name AT %DB930.DBX6198.0, 1 s
   "DB930_Tools_Tool{183}_tool_name" : String[20] = PLC DB930_Tools.Tool[183].tool_name AT %DB930.DBX6232.0, 1 s
   "DB930_Tools_Tool{184}_tool_name" : String[20] = PLC DB930_Tools.Tool[184].tool_name AT %DB930.DBX6266.0, 1 s
   "DB930_Tools_Tool{185}_tool_name" : String[20] = PLC DB930_Tools.Tool[185].tool_name AT %DB930.DBX6300.0, 1 s
   "DB930_Tools_Tool{186}_tool_name" : String[20] = PLC DB930_Tools.Tool[186].tool_name AT %DB930.DBX6334.0, 1 s
   "DB930_Tools_Tool{187}_tool_name" : String[20] = PLC DB930_Tools.Tool[187].tool_name AT %DB930.DBX6368.0, 1 s
   "DB930_Tools_Tool{188}_tool_name" : String[20] = PLC DB930_Tools.Tool[188].tool_name AT %DB930.DBX6402.0, 1 s
   "DB930_Tools_Tool{189}_tool_name" : String[20] = PLC DB930_Tools.Tool[189].tool_name AT %DB930.DBX6436.0, 1 s
   "DB930_Tools_Tool{190}_tool_name" : String[20] = PLC DB930_Tools.Tool[190].tool_name AT %DB930.DBX6470.0, 1 s
   "DB930_Tools_Tool{191}_tool_name" : String[20] = PLC DB930_Tools.Tool[191].tool_name AT %DB930.DBX6504.0, 1 s
   "DB930_Tools_Tool{192}_tool_name" : String[20] = PLC DB930_Tools.Tool[192].tool_name AT %DB930.DBX6538.0, 1 s
   "DB930_Tools_Tool{193}_tool_name" : String[20] = PLC DB930_Tools.Tool[193].tool_name AT %DB930.DBX6572.0, 1 s
   "DB930_Tools_Tool{194}_tool_name" : String[20] = PLC DB930_Tools.Tool[194].tool_name AT %DB930.DBX6606.0, 1 s
   "DB930_Tools_Tool{195}_tool_name" : String[20] = PLC DB930_Tools.Tool[195].tool_name AT %DB930.DBX6640.0, 1 s
   "DB930_Tools_Tool{196}_tool_name" : String[20] = PLC DB930_Tools.Tool[196].tool_name AT %DB930.DBX6674.0, 1 s
   "DB930_Tools_Tool{197}_tool_name" : String[20] = PLC DB930_Tools.Tool[197].tool_name AT %DB930.DBX6708.0, 1 s
   "DB930_Tools_Tool{198}_tool_name" : String[20] = PLC DB930_Tools.Tool[198].tool_name AT %DB930.DBX6742.0, 1 s
   "DB930_Tools_Tool{199}_tool_name" : String[20] = PLC DB930_Tools.Tool[199].tool_name AT %DB930.DBX6776.0, 1 s
   "DB930_Tools_Tool{200}_tool_name" : String[20] = PLC DB930_Tools.Tool[200].tool_name AT %DB930.DBX6810.0, 1 s
   "DB_MouldEditor_HMI_uData_sStatusBits" : Int AT %DB10.DBW812, 1 s
   "InterfaceVisu_MaxFlow{1}" : Real = PLC InterfaceVisu.MaxFlow[1] AT %DB1.DBD320, 1 s
   "InterfaceVisu_MaxFlow{2}" : Real = PLC InterfaceVisu.MaxFlow[2] AT %DB1.DBD324, 1 s
   "InterfaceVisu_MaxFlow{3}" : Real = PLC InterfaceVisu.MaxFlow[3] AT %DB1.DBD328, 1 s
   "InterfaceVisu_MaxFlow{4}" : Real = PLC InterfaceVisu.MaxFlow[4] AT %DB1.DBD332, 1 s
   "InterfaceVisu_MaxFlow{5}" : Real = PLC InterfaceVisu.MaxFlow[5] AT %DB1.DBD336, 1 s
   "InterfaceVisu_MaxFlow{6}" : Real = PLC InterfaceVisu.MaxFlow[6] AT %DB1.DBD340, 1 s
   "InterfaceVisu_MaxTotalFlow{1}" : Real = PLC InterfaceVisu.MaxTotalFlow[1] AT %DB1.DBD348, 1 s
   "InterfaceVisu_MaxTotalFlow{2}" : Real = PLC InterfaceVisu.MaxTotalFlow[2] AT %DB1.DBD352, 1 s
   "InterfaceVisu_MaxTotalFlow{3}" : Real = PLC InterfaceVisu.MaxTotalFlow[3] AT %DB1.DBD356, 1 s
   "InterfaceVisu_MaxTotalFlow{4}" : Real = PLC InterfaceVisu.MaxTotalFlow[4] AT %DB1.DBD360, 1 s
   "InterfaceVisu_MaxTotalFlow{5}" : Real = PLC InterfaceVisu.MaxTotalFlow[5] AT %DB1.DBD364, 1 s
   "InterfaceVisu_MaxTotalFlow{6}" : Real = PLC InterfaceVisu.MaxTotalFlow[6] AT %DB1.DBD368, 1 s
   "InterfaceVisu_MaxTotalFlow{7}" : Real = PLC InterfaceVisu.MaxTotalFlow[7] AT %DB1.DBD372, 1 s
   "InterfaceVisu_MaxTotalFlow{8}" : Real = PLC InterfaceVisu.MaxTotalFlow[8] AT %DB1.DBD376, 1 s
   "InterfaceVisu_MinFlow{1}" : Real = PLC InterfaceVisu.MinFlow[1] AT %DB1.DBD296, 1 s
   "InterfaceVisu_MinFlow{2}" : Real = PLC InterfaceVisu.MinFlow[2] AT %DB1.DBD300, 1 s
   "InterfaceVisu_MinFlow{3}" : Real = PLC InterfaceVisu.MinFlow[3] AT %DB1.DBD304, 1 s
   "InterfaceVisu_MinFlow{4}" : Real = PLC InterfaceVisu.MinFlow[4] AT %DB1.DBD308, 1 s
   "InterfaceVisu_MinFlow{5}" : Real = PLC InterfaceVisu.MinFlow[5] AT %DB1.DBD312, 1 s
   "InterfaceVisu_MinFlow{6}" : Real = PLC InterfaceVisu.MinFlow[6] AT %DB1.DBD316, 1 s
   "InterfaceVisu_HPValuesSet" : Bool = PLC InterfaceVisu.HPValuesSet AT %DB1.DBX104.6, 1 s

